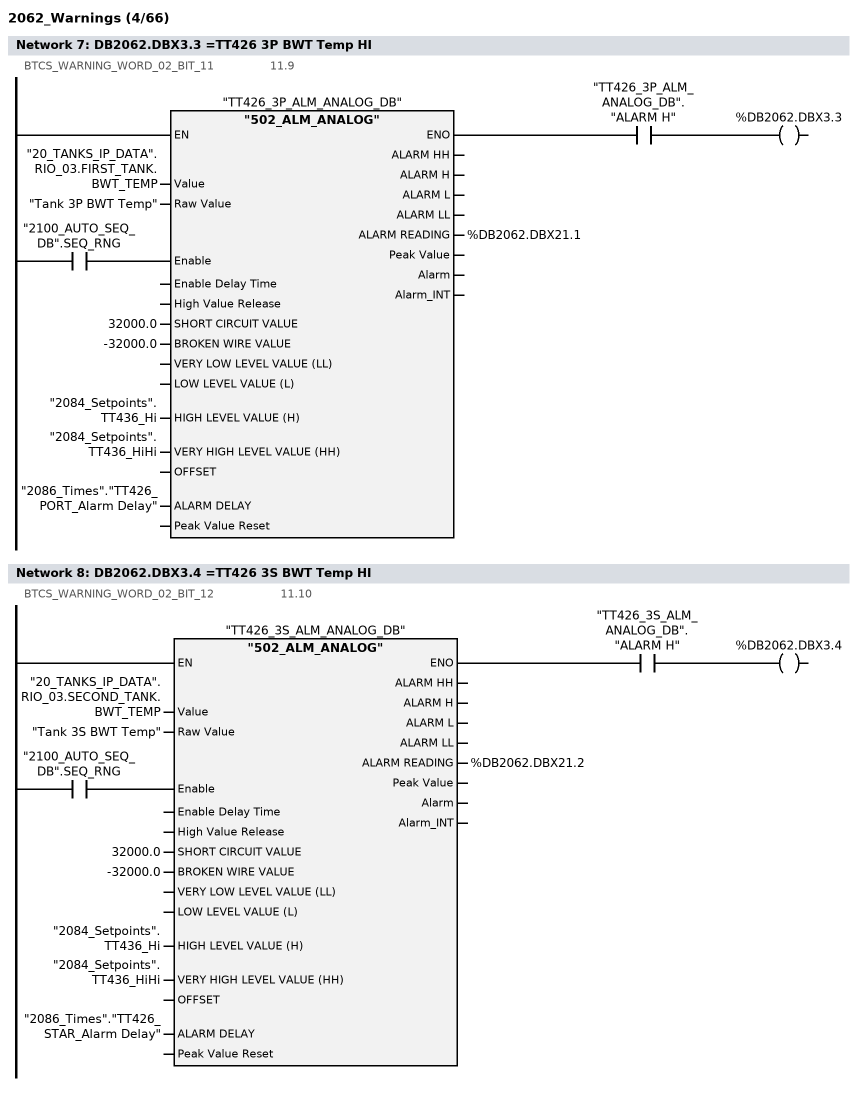
   RUNG wire#powerrail
      "TT426_3P_ALM_ANALOG_DB"(Enable := wire#w1, Value := "20_TANKS_IP_DATA".RIO_03.FIRST_TANK.BWT_TEMP, "Raw Value" := "Tank 3P BWT Temp", "Enable Delay Time" :=, "High Value Release" :=, "SHORT CIRCUIT VALUE" := 32000.0, "BROKEN WIRE VALUE" := -32000.0, "VERY LOW LEVEL VALUE (LL)" :=, "LOW LEVEL VALUE (L)" :=, "HIGH LEVEL VALUE (H)" := "2084_Setpoints".TT436_Hi, "VERY HIGH LEVEL VALUE (HH)" := "2084_Setpoints".TT436_HiHi, OFFSET :=, "ALARM DELAY" := "2086_Times"."TT426_PORT_Alarm Delay", "Peak Value Reset" :=, "ALARM HH" =>, "ALARM H" =>, "ALARM L" =>, "ALARM LL" =>, "ALARM READING" => %DB2062.DBX21.1, "Peak Value" =>, Alarm =>, Alarm_INT =>)
      Contact( "TT426_3P_ALM_ANALOG_DB"."ALARM H" )
      Coil( %DB2062.DBX3.3 )
   END_RUNG
   RUNG wire#powerrail
      Contact( "2100_AUTO_SEQ_DB".SEQ_RNG )
   END_RUNG wire#w1
   // the same network as SCL:
   "TT426_3P_ALM_ANALOG_DB"(Value := "20_TANKS_IP_DATA".RIO_03.FIRST_TANK.BWT_TEMP,   // "502_ALM_ANALOG"
                           "Raw Value" := "Tank 3P BWT Temp",
                           Enable := "2100_AUTO_SEQ_DB".SEQ_RNG,
                           "SHORT CIRCUIT VALUE" := 32000.0,
                           "BROKEN WIRE VALUE" := -32000.0,
                           "HIGH LEVEL VALUE (H)" := "2084_Setpoints".TT436_Hi,
                           "VERY HIGH LEVEL VALUE (HH)" := "2084_Setpoints".TT436_HiHi,
                           "ALARM DELAY" := "2086_Times"."TT426_PORT_Alarm Delay",
                           "ALARM READING" => %DB2062.DBX21.1,
                           ENO => #_w1);
   %DB2062.DBX3.3 := #_w1 AND "TT426_3P_ALM_ANALOG_DB"."ALARM H";
END_REGION

REGION Network 8: DB2062.DBX3.4 =TT426 3S BWT Temp HI
   // BTCS_WARNING_WORD_02_BIT_12                   11.10
   RUNG wire#powerrail
      "TT426_3S_ALM_ANALOG_DB"(Enable := wire#w1, Value := "20_TANKS_IP_DATA".RIO_03.SECOND_TANK.BWT_TEMP, "Raw Value" := "Tank 3S BWT Temp", "Enable Delay Time" :=, "High Value Release" :=, "SHORT CIRCUIT VALUE" := 32000.0, "BROKEN WIRE VALUE" := -32000.0, "VERY LOW LEVEL VALUE (LL)" :=, "LOW LEVEL VALUE (L)" :=, "HIGH LEVEL VALUE (H)" := "2084_Setpoints".TT436_Hi, "VERY HIGH LEVEL VALUE (HH)" := "2084_Setpoints".TT436_HiHi, OFFSET :=, "ALARM DELAY" := "2086_Times"."TT426_STAR_Alarm Delay", "Peak Value Reset" :=, "ALARM HH" =>, "ALARM H" =>, "ALARM L" =>, "ALARM LL" =>, "ALARM READING" => %DB2062.DBX21.2, "Peak Value" =>, Alarm =>, Alarm_INT =>)
      Contact( "TT426_3S_ALM_ANALOG_DB"."ALARM H" )
      Coil( %DB2062.DBX3.4 )
   END_RUNG
   RUNG wire#powerrail
      Contact( "2100_AUTO_SEQ_DB".SEQ_RNG )
   END_RUNG wire#w1
   // the same network as SCL:
   "TT426_3S_ALM_ANALOG_DB"(Value := "20_TANKS_IP_DATA".RIO_03.SECOND_TANK.BWT_TEMP,   // "502_ALM_ANALOG"
                           "Raw Value" := "Tank 3S BWT Temp",
                           Enable := "2100_AUTO_SEQ_DB".SEQ_RNG,
                           "SHORT CIRCUIT VALUE" := 32000.0,
                           "BROKEN WIRE VALUE" := -32000.0,
                           "HIGH LEVEL VALUE (H)" := "2084_Setpoints".TT436_Hi,
                           "VERY HIGH LEVEL VALUE (HH)" := "2084_Setpoints".TT436_HiHi,
                           "ALARM DELAY" := "2086_Times"."TT426_STAR_Alarm Delay",
                           "ALARM READING" => %DB2062.DBX21.2,
                           ENO => #_w1);
   %DB2062.DBX3.4 := #_w1 AND "TT426_3S_ALM_ANALOG_DB"."ALARM H";
END_REGION

REGION Network 9: DB2062.DBX3.5 =TT426 4P BWT Temp HI
   // BTCS_WARNING_WORD_02_BIT_13                     11.11
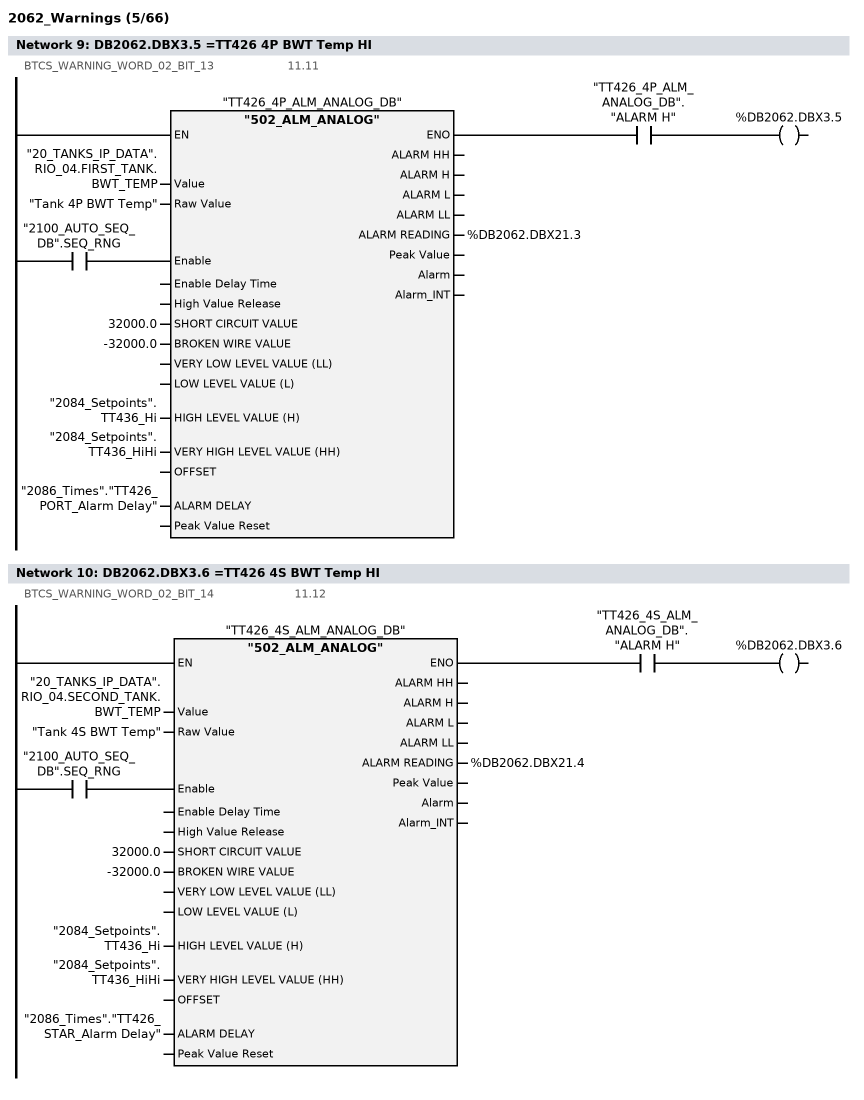
   RUNG wire#powerrail
      "TT426_4P_ALM_ANALOG_DB"(Enable := wire#w1, Value := "20_TANKS_IP_DATA".RIO_04.FIRST_TANK.BWT_TEMP, "Raw Value" := "Tank 4P BWT Temp", "Enable Delay Time" :=, "High Value Release" :=, "SHORT CIRCUIT VALUE" := 32000.0, "BROKEN WIRE VALUE" := -32000.0, "VERY LOW LEVEL VALUE (LL)" :=, "LOW LEVEL VALUE (L)" :=, "HIGH LEVEL VALUE (H)" := "2084_Setpoints".TT436_Hi, "VERY HIGH LEVEL VALUE (HH)" := "2084_Setpoints".TT436_HiHi, OFFSET :=, "ALARM DELAY" := "2086_Times"."TT426_PORT_Alarm Delay", "Peak Value Reset" :=, "ALARM HH" =>, "ALARM H" =>, "ALARM L" =>, "ALARM LL" =>, "ALARM READING" => %DB2062.DBX21.3, "Peak Value" =>, Alarm =>, Alarm_INT =>)
      Contact( "TT426_4P_ALM_ANALOG_DB"."ALARM H" )
      Coil( %DB2062.DBX3.5 )
   END_RUNG
   RUNG wire#powerrail
      Contact( "2100_AUTO_SEQ_DB".SEQ_RNG )
   END_RUNG wire#w1
   // the same network as SCL:
   "TT426_4P_ALM_ANALOG_DB"(Value := "20_TANKS_IP_DATA".RIO_04.FIRST_TANK.BWT_TEMP,   // "502_ALM_ANALOG"
                           "Raw Value" := "Tank 4P BWT Temp",
                           Enable := "2100_AUTO_SEQ_DB".SEQ_RNG,
                           "SHORT CIRCUIT VALUE" := 32000.0,
                           "BROKEN WIRE VALUE" := -32000.0,
                           "HIGH LEVEL VALUE (H)" := "2084_Setpoints".TT436_Hi,
                           "VERY HIGH LEVEL VALUE (HH)" := "2084_Setpoints".TT436_HiHi,
                           "ALARM DELAY" := "2086_Times"."TT426_PORT_Alarm Delay",
                           "ALARM READING" => %DB2062.DBX21.3,
                           ENO => #_w1);
   %DB2062.DBX3.5 := #_w1 AND "TT426_4P_ALM_ANALOG_DB"."ALARM H";
END_REGION

REGION Network 10: DB2062.DBX3.6 =TT426 4S BWT Temp HI
   // BTCS_WARNING_WORD_02_BIT_14                       11.12
   RUNG wire#powerrail
      "TT426_4S_ALM_ANALOG_DB"(Enable := wire#w1, Value := "20_TANKS_IP_DATA".RIO_04.SECOND_TANK.BWT_TEMP, "Raw Value" := "Tank 4S BWT Temp", "Enable Delay Time" :=, "High Value Release" :=, "SHORT CIRCUIT VALUE" := 32000.0, "BROKEN WIRE VALUE" := -32000.0, "VERY LOW LEVEL VALUE (LL)" :=, "LOW LEVEL VALUE (L)" :=, "HIGH LEVEL VALUE (H)" := "2084_Setpoints".TT436_Hi, "VERY HIGH LEVEL VALUE (HH)" := "2084_Setpoints".TT436_HiHi, OFFSET :=, "ALARM DELAY" := "2086_Times"."TT426_STAR_Alarm Delay", "Peak Value Reset" :=, "ALARM HH" =>, "ALARM H" =>, "ALARM L" =>, "ALARM LL" =>, "ALARM READING" => %DB2062.DBX21.4, "Peak Value" =>, Alarm =>, Alarm_INT =>)
      Contact( "TT426_4S_ALM_ANALOG_DB"."ALARM H" )
      Coil( %DB2062.DBX3.6 )
   END_RUNG
   RUNG wire#powerrail
      Contact( "2100_AUTO_SEQ_DB".SEQ_RNG )
   END_RUNG wire#w1
   // the same network as SCL:
   "TT426_4S_ALM_ANALOG_DB"(Value := "20_TANKS_IP_DATA".RIO_04.SECOND_TANK.BWT_TEMP,   // "502_ALM_ANALOG"
                           "Raw Value" := "Tank 4S BWT Temp",
                           Enable := "2100_AUTO_SEQ_DB".SEQ_RNG,
                           "SHORT CIRCUIT VALUE" := 32000.0,
                           "BROKEN WIRE VALUE" := -32000.0,
                           "HIGH LEVEL VALUE (H)" := "2084_Setpoints".TT436_Hi,
                           "VERY HIGH LEVEL VALUE (HH)" := "2084_Setpoints".TT436_HiHi,
                           "ALARM DELAY" := "2086_Times"."TT426_STAR_Alarm Delay",
                           "ALARM READING" => %DB2062.DBX21.4,
                           ENO => #_w1);
   %DB2062.DBX3.6 := #_w1 AND "TT426_4S_ALM_ANALOG_DB"."ALARM H";
END_REGION

REGION Network 11: DB2062.DBX3.7 =TT426 5P BWT Temp HI
   // BTCS_WARNING_WORD_02_BIT_15                        11.13
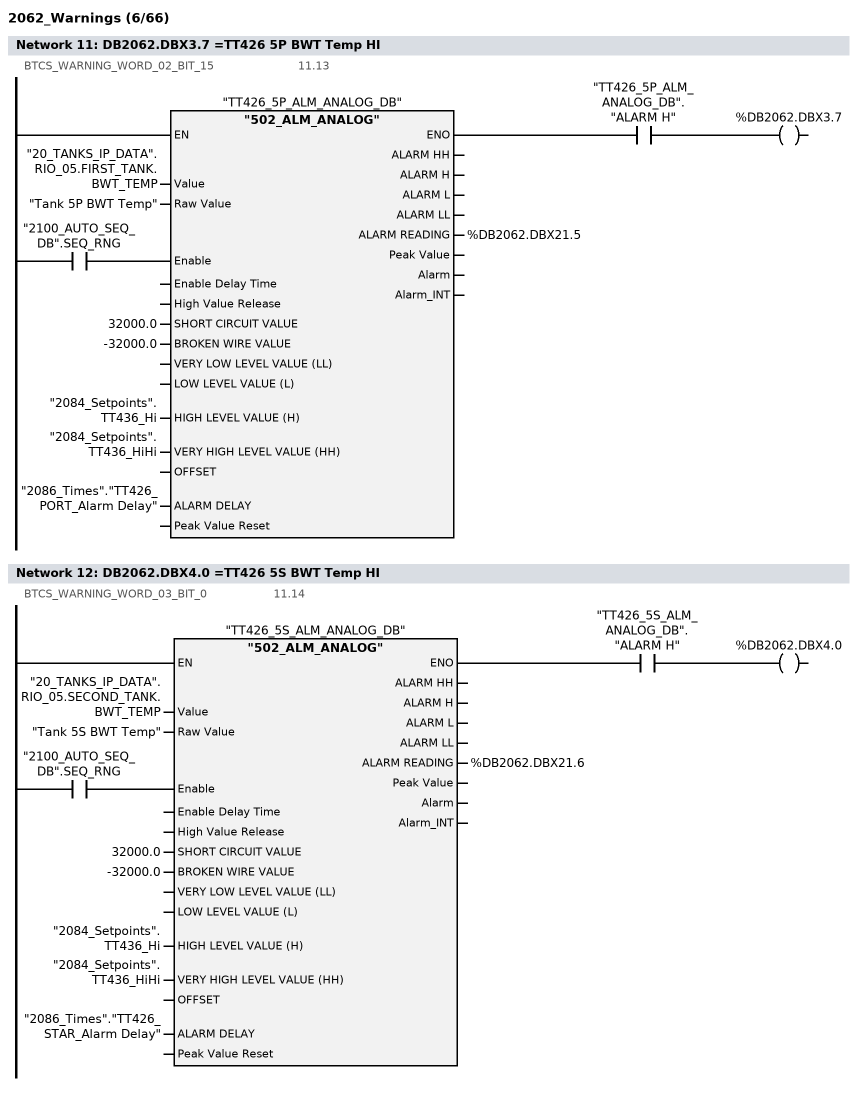
   RUNG wire#powerrail
      "TT426_5P_ALM_ANALOG_DB"(Enable := wire#w1, Value := "20_TANKS_IP_DATA".RIO_05.FIRST_TANK.BWT_TEMP, "Raw Value" := "Tank 5P BWT Temp", "Enable Delay Time" :=, "High Value Release" :=, "SHORT CIRCUIT VALUE" := 32000.0, "BROKEN WIRE VALUE" := -32000.0, "VERY LOW LEVEL VALUE (LL)" :=, "LOW LEVEL VALUE (L)" :=, "HIGH LEVEL VALUE (H)" := "2084_Setpoints".TT436_Hi, "VERY HIGH LEVEL VALUE (HH)" := "2084_Setpoints".TT436_HiHi, OFFSET :=, "ALARM DELAY" := "2086_Times"."TT426_PORT_Alarm Delay", "Peak Value Reset" :=, "ALARM HH" =>, "ALARM H" =>, "ALARM L" =>, "ALARM LL" =>, "ALARM READING" => %DB2062.DBX21.5, "Peak Value" =>, Alarm =>, Alarm_INT =>)
      Contact( "TT426_5P_ALM_ANALOG_DB"."ALARM H" )
      Coil( %DB2062.DBX3.7 )
   END_RUNG
   RUNG wire#powerrail
      Contact( "2100_AUTO_SEQ_DB".SEQ_RNG )
   END_RUNG wire#w1
   // the same network as SCL:
   "TT426_5P_ALM_ANALOG_DB"(Value := "20_TANKS_IP_DATA".RIO_05.FIRST_TANK.BWT_TEMP,   // "502_ALM_ANALOG"
                           "Raw Value" := "Tank 5P BWT Temp",
                           Enable := "2100_AUTO_SEQ_DB".SEQ_RNG,
                           "SHORT CIRCUIT VALUE" := 32000.0,
                           "BROKEN WIRE VALUE" := -32000.0,
                           "HIGH LEVEL VALUE (H)" := "2084_Setpoints".TT436_Hi,
                           "VERY HIGH LEVEL VALUE (HH)" := "2084_Setpoints".TT436_HiHi,
                           "ALARM DELAY" := "2086_Times"."TT426_PORT_Alarm Delay",
                           "ALARM READING" => %DB2062.DBX21.5,
                           ENO => #_w1);
   %DB2062.DBX3.7 := #_w1 AND "TT426_5P_ALM_ANALOG_DB"."ALARM H";
END_REGION

REGION Network 12: DB2062.DBX4.0 =TT426 5S BWT Temp HI
   // BTCS_WARNING_WORD_03_BIT_0                   11.14
   RUNG wire#powerrail
      "TT426_5S_ALM_ANALOG_DB"(Enable := wire#w1, Value := "20_TANKS_IP_DATA".RIO_05.SECOND_TANK.BWT_TEMP, "Raw Value" := "Tank 5S BWT Temp", "Enable Delay Time" :=, "High Value Release" :=, "SHORT CIRCUIT VALUE" := 32000.0, "BROKEN WIRE VALUE" := -32000.0, "VERY LOW LEVEL VALUE (LL)" :=, "LOW LEVEL VALUE (L)" :=, "HIGH LEVEL VALUE (H)" := "2084_Setpoints".TT436_Hi, "VERY HIGH LEVEL VALUE (HH)" := "2084_Setpoints".TT436_HiHi, OFFSET :=, "ALARM DELAY" := "2086_Times"."TT426_STAR_Alarm Delay", "Peak Value Reset" :=, "ALARM HH" =>, "ALARM H" =>, "ALARM L" =>, "ALARM LL" =>, "ALARM READING" => %DB2062.DBX21.6, "Peak Value" =>, Alarm =>, Alarm_INT =>)
      Contact( "TT426_5S_ALM_ANALOG_DB"."ALARM H" )
      Coil( %DB2062.DBX4.0 )
   END_RUNG
   RUNG wire#powerrail
      Contact( "2100_AUTO_SEQ_DB".SEQ_RNG )
   END_RUNG wire#w1
   // the same network as SCL:
   "TT426_5S_ALM_ANALOG_DB"(Value := "20_TANKS_IP_DATA".RIO_05.SECOND_TANK.BWT_TEMP,   // "502_ALM_ANALOG"
                           "Raw Value" := "Tank 5S BWT Temp",
                           Enable := "2100_AUTO_SEQ_DB".SEQ_RNG,
                           "SHORT CIRCUIT VALUE" := 32000.0,
                           "BROKEN WIRE VALUE" := -32000.0,
                           "HIGH LEVEL VALUE (H)" := "2084_Setpoints".TT436_Hi,
                           "VERY HIGH LEVEL VALUE (HH)" := "2084_Setpoints".TT436_HiHi,
                           "ALARM DELAY" := "2086_Times"."TT426_STAR_Alarm Delay",
                           "ALARM READING" => %DB2062.DBX21.6,
                           ENO => #_w1);
   %DB2062.DBX4.0 := #_w1 AND "TT426_5S_ALM_ANALOG_DB"."ALARM H";
END_REGION

REGION Network 13: DB2062.DBX4.1 =TT426 6P BWT Temp HI
   // BTCS_WARNING_WORD_03_BIT_1                           11.15
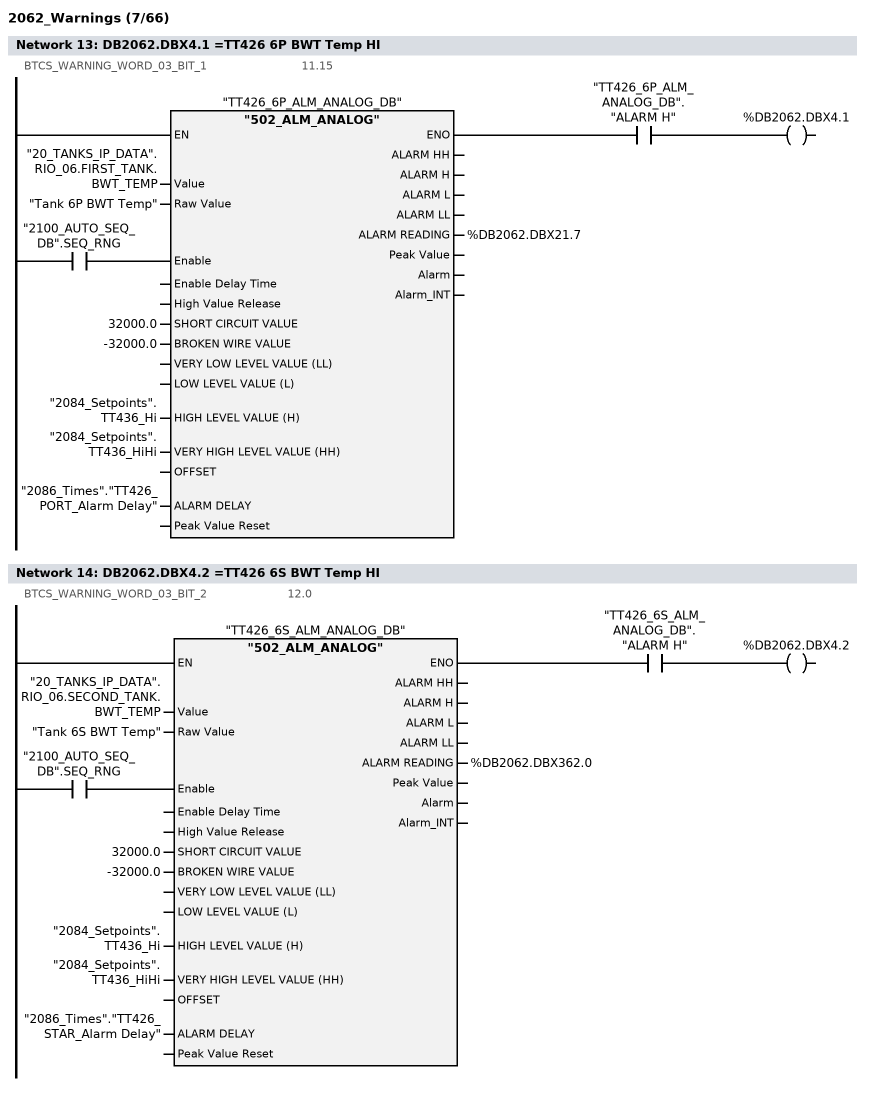
   RUNG wire#powerrail
      "TT426_6P_ALM_ANALOG_DB"(Enable := wire#w1, Value := "20_TANKS_IP_DATA".RIO_06.FIRST_TANK.BWT_TEMP, "Raw Value" := "Tank 6P BWT Temp", "Enable Delay Time" :=, "High Value Release" :=, "SHORT CIRCUIT VALUE" := 32000.0, "BROKEN WIRE VALUE" := -32000.0, "VERY LOW LEVEL VALUE (LL)" :=, "LOW LEVEL VALUE (L)" :=, "HIGH LEVEL VALUE (H)" := "2084_Setpoints".TT436_Hi, "VERY HIGH LEVEL VALUE (HH)" := "2084_Setpoints".TT436_HiHi, OFFSET :=, "ALARM DELAY" := "2086_Times"."TT426_PORT_Alarm Delay", "Peak Value Reset" :=, "ALARM HH" =>, "ALARM H" =>, "ALARM L" =>, "ALARM LL" =>, "ALARM READING" => %DB2062.DBX21.7, "Peak Value" =>, Alarm =>, Alarm_INT =>)
      Contact( "TT426_6P_ALM_ANALOG_DB"."ALARM H" )
      Coil( %DB2062.DBX4.1 )
   END_RUNG
   RUNG wire#powerrail
      Contact( "2100_AUTO_SEQ_DB".SEQ_RNG )
   END_RUNG wire#w1
   // the same network as SCL:
   "TT426_6P_ALM_ANALOG_DB"(Value := "20_TANKS_IP_DATA".RIO_06.FIRST_TANK.BWT_TEMP,   // "502_ALM_ANALOG"
                           "Raw Value" := "Tank 6P BWT Temp",
                           Enable := "2100_AUTO_SEQ_DB".SEQ_RNG,
                           "SHORT CIRCUIT VALUE" := 32000.0,
                           "BROKEN WIRE VALUE" := -32000.0,
                           "HIGH LEVEL VALUE (H)" := "2084_Setpoints".TT436_Hi,
                           "VERY HIGH LEVEL VALUE (HH)" := "2084_Setpoints".TT436_HiHi,
                           "ALARM DELAY" := "2086_Times"."TT426_PORT_Alarm Delay",
                           "ALARM READING" => %DB2062.DBX21.7,
                           ENO => #_w1);
   %DB2062.DBX4.1 := #_w1 AND "TT426_6P_ALM_ANALOG_DB"."ALARM H";
END_REGION

REGION Network 14: DB2062.DBX4.2 =TT426 6S BWT Temp HI
   // BTCS_WARNING_WORD_03_BIT_2                       12.0
   RUNG wire#powerrail
      "TT426_6S_ALM_ANALOG_DB"(Enable := wire#w1, Value := "20_TANKS_IP_DATA".RIO_06.SECOND_TANK.BWT_TEMP, "Raw Value" := "Tank 6S BWT Temp", "Enable Delay Time" :=, "High Value Release" :=, "SHORT CIRCUIT VALUE" := 32000.0, "BROKEN WIRE VALUE" := -32000.0, "VERY LOW LEVEL VALUE (LL)" :=, "LOW LEVEL VALUE (L)" :=, "HIGH LEVEL VALUE (H)" := "2084_Setpoints".TT436_Hi, "VERY HIGH LEVEL VALUE (HH)" := "2084_Setpoints".TT436_HiHi, OFFSET :=, "ALARM DELAY" := "2086_Times"."TT426_STAR_Alarm Delay", "Peak Value Reset" :=, "ALARM HH" =>, "ALARM H" =>, "ALARM L" =>, "ALARM LL" =>, "ALARM READING" => %DB2062.DBX362.0, "Peak Value" =>, Alarm =>, Alarm_INT =>)
      Contact( "TT426_6S_ALM_ANALOG_DB"."ALARM H" )
      Coil( %DB2062.DBX4.2 )
   END_RUNG
   RUNG wire#powerrail
      Contact( "2100_AUTO_SEQ_DB".SEQ_RNG )
   END_RUNG wire#w1
   // the same network as SCL:
   "TT426_6S_ALM_ANALOG_DB"(Value := "20_TANKS_IP_DATA".RIO_06.SECOND_TANK.BWT_TEMP,   // "502_ALM_ANALOG"
                           "Raw Value" := "Tank 6S BWT Temp",
                           Enable := "2100_AUTO_SEQ_DB".SEQ_RNG,
                           "SHORT CIRCUIT VALUE" := 32000.0,
                           "BROKEN WIRE VALUE" := -32000.0,
                           "HIGH LEVEL VALUE (H)" := "2084_Setpoints".TT436_Hi,
                           "VERY HIGH LEVEL VALUE (HH)" := "2084_Setpoints".TT436_HiHi,
                           "ALARM DELAY" := "2086_Times"."TT426_STAR_Alarm Delay",
                           "ALARM READING" => %DB2062.DBX362.0,
                           ENO => #_w1);
   %DB2062.DBX4.2 := #_w1 AND "TT426_6S_ALM_ANALOG_DB"."ALARM H";
END_REGION

REGION Network 15: DB2062.DBX4.3 =TT426 APT BWT Temp HI
   // BTCS_WARNING_WORD_03_BIT_3                                 12.1
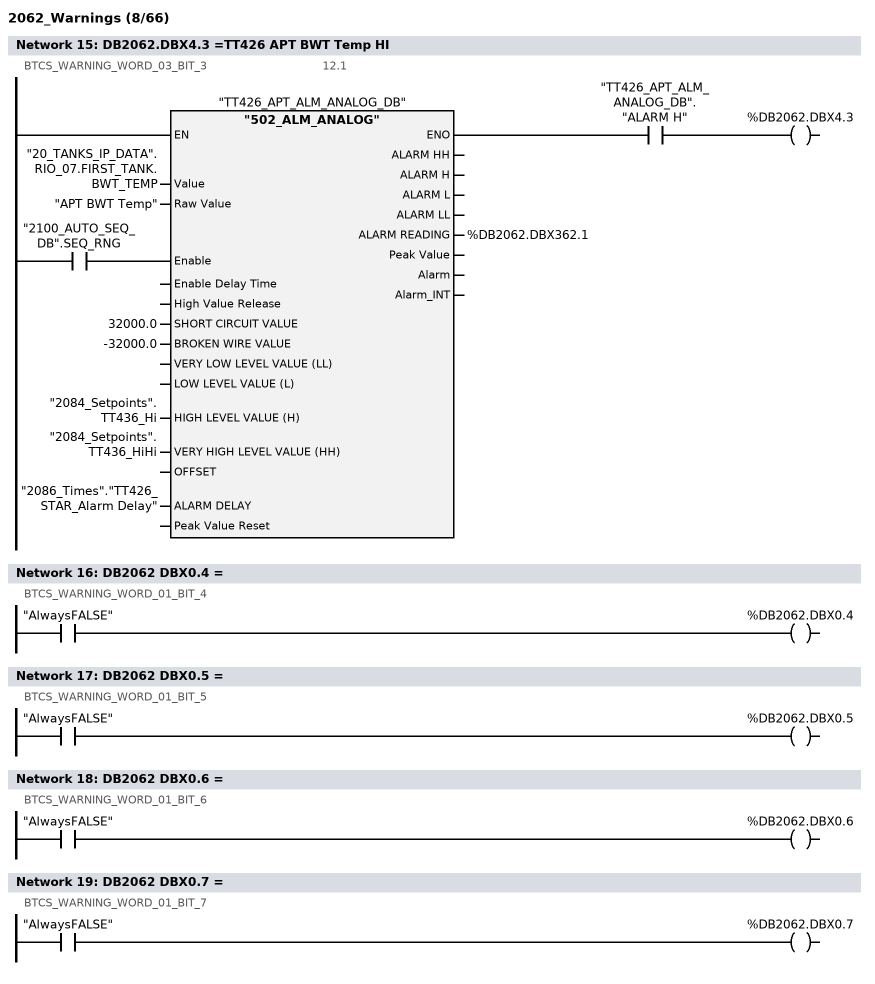
   RUNG wire#powerrail
      "TT426_APT_ALM_ANALOG_DB"(Enable := wire#w1, Value := "20_TANKS_IP_DATA".RIO_07.FIRST_TANK.BWT_TEMP, "Raw Value" := "APT BWT Temp", "Enable Delay Time" :=, "High Value Release" :=, "SHORT CIRCUIT VALUE" := 32000.0, "BROKEN WIRE VALUE" := -32000.0, "VERY LOW LEVEL VALUE (LL)" :=, "LOW LEVEL VALUE (L)" :=, "HIGH LEVEL VALUE (H)" := "2084_Setpoints".TT436_Hi, "VERY HIGH LEVEL VALUE (HH)" := "2084_Setpoints".TT436_HiHi, OFFSET :=, "ALARM DELAY" := "2086_Times"."TT426_STAR_Alarm Delay", "Peak Value Reset" :=, "ALARM HH" =>, "ALARM H" =>, "ALARM L" =>, "ALARM LL" =>, "ALARM READING" => %DB2062.DBX362.1, "Peak Value" =>, Alarm =>, Alarm_INT =>)
      Contact( "TT426_APT_ALM_ANALOG_DB"."ALARM H" )
      Coil( %DB2062.DBX4.3 )
   END_RUNG
   RUNG wire#powerrail
      Contact( "2100_AUTO_SEQ_DB".SEQ_RNG )
   END_RUNG wire#w1
   // the same network as SCL:
   "TT426_APT_ALM_ANALOG_DB"(Value := "20_TANKS_IP_DATA".RIO_07.FIRST_TANK.BWT_TEMP,   // "502_ALM_ANALOG"
                           "Raw Value" := "APT BWT Temp",
                           Enable := "2100_AUTO_SEQ_DB".SEQ_RNG,
                           "SHORT CIRCUIT VALUE" := 32000.0,
                           "BROKEN WIRE VALUE" := -32000.0,
                           "HIGH LEVEL VALUE (H)" := "2084_Setpoints".TT436_Hi,
                           "VERY HIGH LEVEL VALUE (HH)" := "2084_Setpoints".TT436_HiHi,
                           "ALARM DELAY" := "2086_Times"."TT426_STAR_Alarm Delay",
                           "ALARM READING" => %DB2062.DBX362.1,
                           ENO => #_w1);
   %DB2062.DBX4.3 := #_w1 AND "TT426_APT_ALM_ANALOG_DB"."ALARM H";
END_REGION

REGION Network 16: DB2062 DBX0.4 =
   // BTCS_WARNING_WORD_01_BIT_4
   RUNG wire#powerrail
      Contact( "AlwaysFALSE" )
      Coil( %DB2062.DBX0.4 )
   END_RUNG
   // the same network as SCL:
   %DB2062.DBX0.4 := "AlwaysFALSE";
END_REGION

REGION Network 17: DB2062 DBX0.5 =
   // BTCS_WARNING_WORD_01_BIT_5
   RUNG wire#powerrail
      Contact( "AlwaysFALSE" )
      Coil( %DB2062.DBX0.5 )
   END_RUNG
   // the same network as SCL:
   %DB2062.DBX0.5 := "AlwaysFALSE";
END_REGION

REGION Network 18: DB2062 DBX0.6 =
   // BTCS_WARNING_WORD_01_BIT_6
   RUNG wire#powerrail
      Contact( "AlwaysFALSE" )
      Coil( %DB2062.DBX0.6 )
   END_RUNG
   // the same network as SCL:
   %DB2062.DBX0.6 := "AlwaysFALSE";
END_REGION

REGION Network 19: DB2062 DBX0.7 =
   // BTCS_WARNING_WORD_01_BIT_7
   RUNG wire#powerrail
      Contact( "AlwaysFALSE" )
      Coil( %DB2062.DBX0.7 )
   END_RUNG
   // the same network as SCL:
   %DB2062.DBX0.7 := "AlwaysFALSE";
END_REGION

REGION Network 20: DB2062.DBX5.0 = FIT418 FPT USD Flow LO / DB2062.DBX5.1 = FIT418 FPT USD Flow HI
   // BTCS_WARNING_WORD_03_BIT_8/9                    12.2
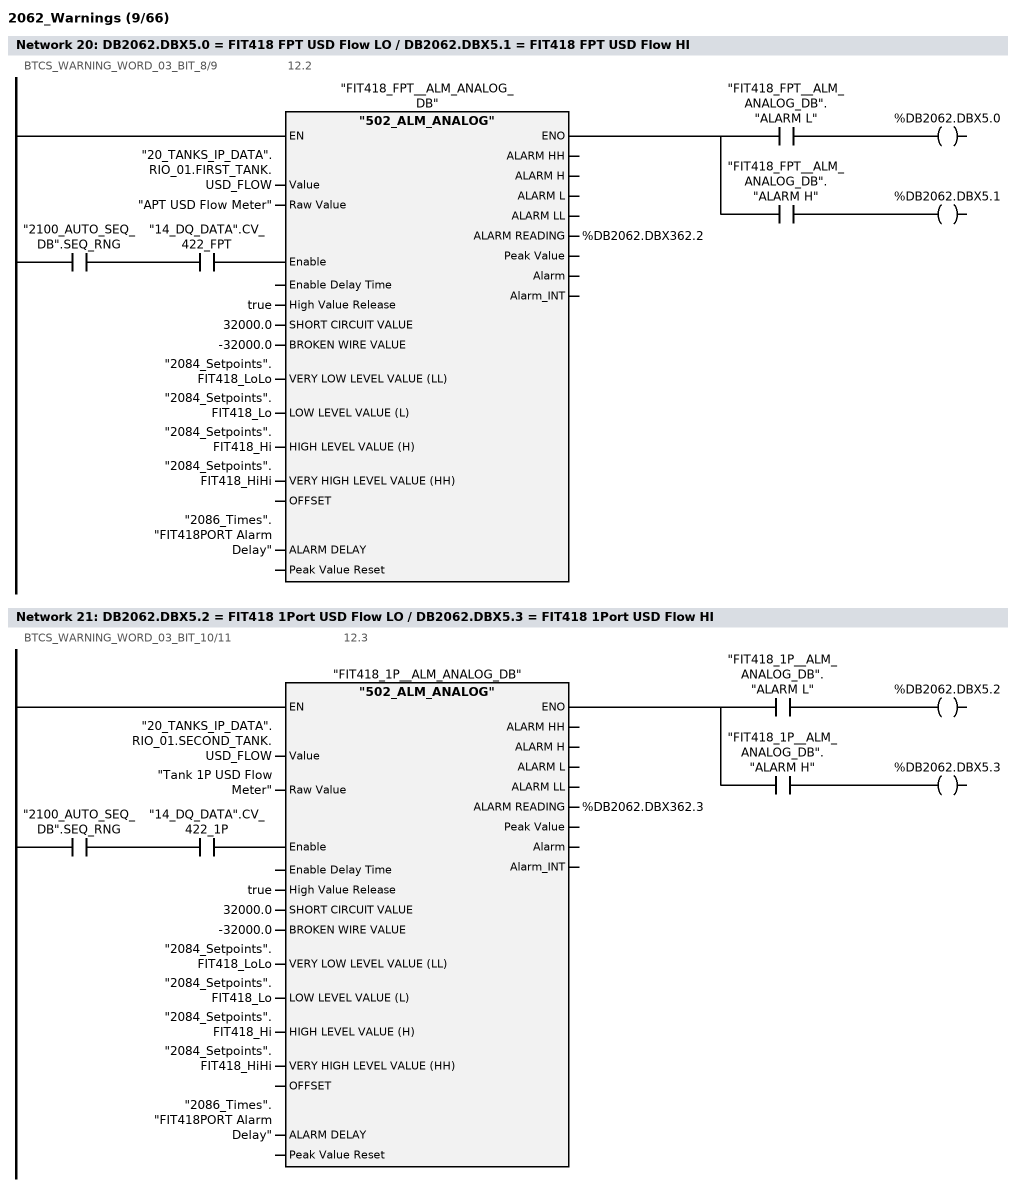
   RUNG wire#powerrail
      "FIT418_FPT__ALM_ANALOG_DB"(Enable := wire#w1, Value := "20_TANKS_IP_DATA".RIO_01.FIRST_TANK.USD_FLOW, "Raw Value" := "APT USD Flow Meter", "Enable Delay Time" :=, "High Value Release" := true, "SHORT CIRCUIT VALUE" := 32000.0, "BROKEN WIRE VALUE" := -32000.0, "VERY LOW LEVEL VALUE (LL)" := "2084_Setpoints".FIT418_LoLo, "LOW LEVEL VALUE (L)" := "2084_Setpoints".FIT418_Lo, "HIGH LEVEL VALUE (H)" := "2084_Setpoints".FIT418_Hi, "VERY HIGH LEVEL VALUE (HH)" := "2084_Setpoints".FIT418_HiHi, OFFSET :=, "ALARM DELAY" := "2086_Times"."FIT418PORT Alarm Delay", "Peak Value Reset" :=, "ALARM HH" =>, "ALARM H" =>, "ALARM L" =>, "ALARM LL" =>, "ALARM READING" => %DB2062.DBX362.2, "Peak Value" =>, Alarm =>, Alarm_INT =>)
      wire#w2
      Contact( "FIT418_FPT__ALM_ANALOG_DB"."ALARM L" )
      Coil( %DB2062.DBX5.0 )
   END_RUNG
   RUNG wire#powerrail
      Contact( "2100_AUTO_SEQ_DB".SEQ_RNG )
      Contact( "14_DQ_DATA".CV_422_FPT )
   END_RUNG wire#w1
   RUNG wire#w2
      Contact( "FIT418_FPT__ALM_ANALOG_DB"."ALARM H" )
      Coil( %DB2062.DBX5.1 )
   END_RUNG
   // the same network as SCL:
   "FIT418_FPT__ALM_ANALOG_DB"(Value := "20_TANKS_IP_DATA".RIO_01.FIRST_TANK.USD_FLOW,   // "502_ALM_ANALOG"
                           "Raw Value" := "APT USD Flow Meter",
                           Enable := "2100_AUTO_SEQ_DB".SEQ_RNG AND "14_DQ_DATA".CV_422_FPT,
                           "High Value Release" := true,
                           "SHORT CIRCUIT VALUE" := 32000.0,
                           "BROKEN WIRE VALUE" := -32000.0,
                           "VERY LOW LEVEL VALUE (LL)" := "2084_Setpoints".FIT418_LoLo,
                           "LOW LEVEL VALUE (L)" := "2084_Setpoints".FIT418_Lo,
                           "HIGH LEVEL VALUE (H)" := "2084_Setpoints".FIT418_Hi,
                           "VERY HIGH LEVEL VALUE (HH)" := "2084_Setpoints".FIT418_HiHi,
                           "ALARM DELAY" := "2086_Times"."FIT418PORT Alarm Delay",
                           "ALARM READING" => %DB2062.DBX362.2,
                           ENO => #_w1);
   %DB2062.DBX5.0 := #_w1 AND "FIT418_FPT__ALM_ANALOG_DB"."ALARM L";
   %DB2062.DBX5.1 := #_w1 AND "FIT418_FPT__ALM_ANALOG_DB"."ALARM H";
END_REGION

REGION Network 21: DB2062.DBX5.2 = FIT418 1Port USD Flow LO / DB2062.DBX5.3 = FIT418 1Port USD Flow HI
   // BTCS_WARNING_WORD_03_BIT_10/11                                12.3
   RUNG wire#powerrail
      "FIT418_1P__ALM_ANALOG_DB"(Enable := wire#w1, Value := "20_TANKS_IP_DATA".RIO_01.SECOND_TANK.USD_FLOW, "Raw Value" := "Tank 1P USD Flow Meter", "Enable Delay Time" :=, "High Value Release" := true, "SHORT CIRCUIT VALUE" := 32000.0, "BROKEN WIRE VALUE" := -32000.0, "VERY LOW LEVEL VALUE (LL)" := "2084_Setpoints".FIT418_LoLo, "LOW LEVEL VALUE (L)" := "2084_Setpoints".FIT418_Lo, "HIGH LEVEL VALUE (H)" := "2084_Setpoints".FIT418_Hi, "VERY HIGH LEVEL VALUE (HH)" := "2084_Setpoints".FIT418_HiHi, OFFSET :=, "ALARM DELAY" := "2086_Times"."FIT418PORT Alarm Delay", "Peak Value Reset" :=, "ALARM HH" =>, "ALARM H" =>, "ALARM L" =>, "ALARM LL" =>, "ALARM READING" => %DB2062.DBX362.3, "Peak Value" =>, Alarm =>, Alarm_INT =>)
      wire#w2
      Contact( "FIT418_1P__ALM_ANALOG_DB"."ALARM L" )
      Coil( %DB2062.DBX5.2 )
   END_RUNG
   RUNG wire#powerrail
      Contact( "2100_AUTO_SEQ_DB".SEQ_RNG )
      Contact( "14_DQ_DATA".CV_422_1P )
   END_RUNG wire#w1
   RUNG wire#w2
      Contact( "FIT418_1P__ALM_ANALOG_DB"."ALARM H" )
      Coil( %DB2062.DBX5.3 )
   END_RUNG
   // the same network as SCL:
   "FIT418_1P__ALM_ANALOG_DB"(Value := "20_TANKS_IP_DATA".RIO_01.SECOND_TANK.USD_FLOW,   // "502_ALM_ANALOG"
                           "Raw Value" := "Tank 1P USD Flow Meter",
                           Enable := "2100_AUTO_SEQ_DB".SEQ_RNG AND "14_DQ_DATA".CV_422_1P,
                           "High Value Release" := true,
                           "SHORT CIRCUIT VALUE" := 32000.0,
                           "BROKEN WIRE VALUE" := -32000.0,
                           "VERY LOW LEVEL VALUE (LL)" := "2084_Setpoints".FIT418_LoLo,
                           "LOW LEVEL VALUE (L)" := "2084_Setpoints".FIT418_Lo,
                           "HIGH LEVEL VALUE (H)" := "2084_Setpoints".FIT418_Hi,
                           "VERY HIGH LEVEL VALUE (HH)" := "2084_Setpoints".FIT418_HiHi,
                           "ALARM DELAY" := "2086_Times"."FIT418PORT Alarm Delay",
                           "ALARM READING" => %DB2062.DBX362.3,
                           ENO => #_w1);
   %DB2062.DBX5.2 := #_w1 AND "FIT418_1P__ALM_ANALOG_DB"."ALARM L";
   %DB2062.DBX5.3 := #_w1 AND "FIT418_1P__ALM_ANALOG_DB"."ALARM H";
END_REGION

REGION Network 22: DB2062.DBX5.4 = FIT417 1Star USD Flow LO / DB2062.DBX5.5 = FIT417 1Star USD Flow HI
   // BTCS_WARNING_WORD_03_BIT_12/13                        12.4
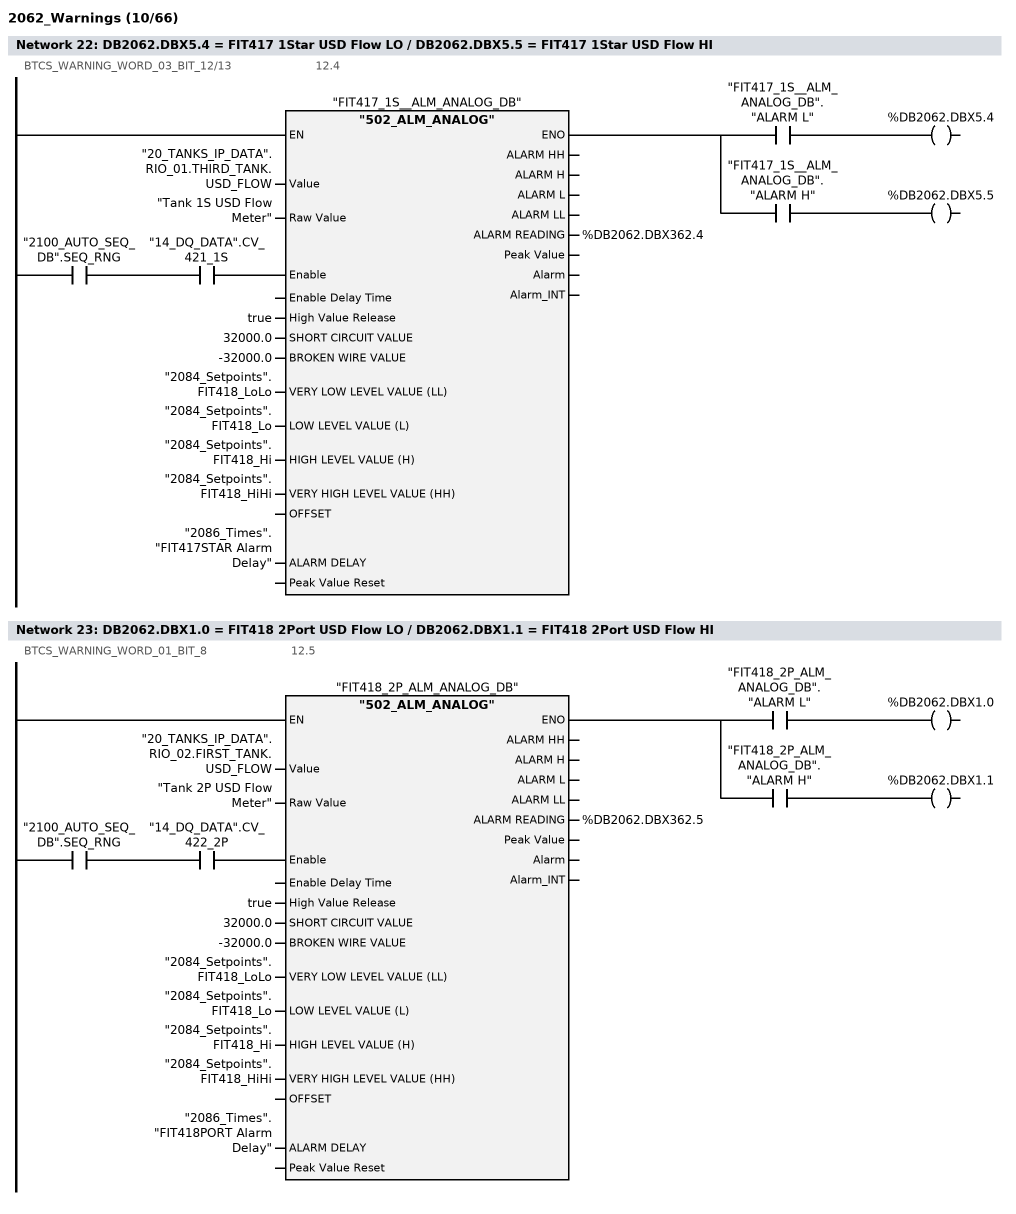
   RUNG wire#powerrail
      "FIT417_1S__ALM_ANALOG_DB"(Enable := wire#w1, Value := "20_TANKS_IP_DATA".RIO_01.THIRD_TANK.USD_FLOW, "Raw Value" := "Tank 1S USD Flow Meter", "Enable Delay Time" :=, "High Value Release" := true, "SHORT CIRCUIT VALUE" := 32000.0, "BROKEN WIRE VALUE" := -32000.0, "VERY LOW LEVEL VALUE (LL)" := "2084_Setpoints".FIT418_LoLo, "LOW LEVEL VALUE (L)" := "2084_Setpoints".FIT418_Lo, "HIGH LEVEL VALUE (H)" := "2084_Setpoints".FIT418_Hi, "VERY HIGH LEVEL VALUE (HH)" := "2084_Setpoints".FIT418_HiHi, OFFSET :=, "ALARM DELAY" := "2086_Times"."FIT417STAR Alarm Delay", "Peak Value Reset" :=, "ALARM HH" =>, "ALARM H" =>, "ALARM L" =>, "ALARM LL" =>, "ALARM READING" => %DB2062.DBX362.4, "Peak Value" =>, Alarm =>, Alarm_INT =>)
      wire#w2
      Contact( "FIT417_1S__ALM_ANALOG_DB"."ALARM L" )
      Coil( %DB2062.DBX5.4 )
   END_RUNG
   RUNG wire#powerrail
      Contact( "2100_AUTO_SEQ_DB".SEQ_RNG )
      Contact( "14_DQ_DATA".CV_421_1S )
   END_RUNG wire#w1
   RUNG wire#w2
      Contact( "FIT417_1S__ALM_ANALOG_DB"."ALARM H" )
      Coil( %DB2062.DBX5.5 )
   END_RUNG
   // the same network as SCL:
   "FIT417_1S__ALM_ANALOG_DB"(Value := "20_TANKS_IP_DATA".RIO_01.THIRD_TANK.USD_FLOW,   // "502_ALM_ANALOG"
                           "Raw Value" := "Tank 1S USD Flow Meter",
                           Enable := "2100_AUTO_SEQ_DB".SEQ_RNG AND "14_DQ_DATA".CV_421_1S,
                           "High Value Release" := true,
                           "SHORT CIRCUIT VALUE" := 32000.0,
                           "BROKEN WIRE VALUE" := -32000.0,
                           "VERY LOW LEVEL VALUE (LL)" := "2084_Setpoints".FIT418_LoLo,
                           "LOW LEVEL VALUE (L)" := "2084_Setpoints".FIT418_Lo,
                           "HIGH LEVEL VALUE (H)" := "2084_Setpoints".FIT418_Hi,
                           "VERY HIGH LEVEL VALUE (HH)" := "2084_Setpoints".FIT418_HiHi,
                           "ALARM DELAY" := "2086_Times"."FIT417STAR Alarm Delay",
                           "ALARM READING" => %DB2062.DBX362.4,
                           ENO => #_w1);
   %DB2062.DBX5.4 := #_w1 AND "FIT417_1S__ALM_ANALOG_DB"."ALARM L";
   %DB2062.DBX5.5 := #_w1 AND "FIT417_1S__ALM_ANALOG_DB"."ALARM H";
END_REGION

REGION Network 23: DB2062.DBX1.0 = FIT418 2Port USD Flow LO / DB2062.DBX1.1 = FIT418 2Port USD Flow HI
   // BTCS_WARNING_WORD_01_BIT_8                        12.5
   RUNG wire#powerrail
      "FIT418_2P_ALM_ANALOG_DB"(Enable := wire#w1, Value := "20_TANKS_IP_DATA".RIO_02.FIRST_TANK.USD_FLOW, "Raw Value" := "Tank 2P USD Flow Meter", "Enable Delay Time" :=, "High Value Release" := true, "SHORT CIRCUIT VALUE" := 32000.0, "BROKEN WIRE VALUE" := -32000.0, "VERY LOW LEVEL VALUE (LL)" := "2084_Setpoints".FIT418_LoLo, "LOW LEVEL VALUE (L)" := "2084_Setpoints".FIT418_Lo, "HIGH LEVEL VALUE (H)" := "2084_Setpoints".FIT418_Hi, "VERY HIGH LEVEL VALUE (HH)" := "2084_Setpoints".FIT418_HiHi, OFFSET :=, "ALARM DELAY" := "2086_Times"."FIT418PORT Alarm Delay", "Peak Value Reset" :=, "ALARM HH" =>, "ALARM H" =>, "ALARM L" =>, "ALARM LL" =>, "ALARM READING" => %DB2062.DBX362.5, "Peak Value" =>, Alarm =>, Alarm_INT =>)
      wire#w2
      Contact( "FIT418_2P_ALM_ANALOG_DB"."ALARM L" )
      Coil( %DB2062.DBX1.0 )
   END_RUNG
   RUNG wire#powerrail
      Contact( "2100_AUTO_SEQ_DB".SEQ_RNG )
      Contact( "14_DQ_DATA".CV_422_2P )
   END_RUNG wire#w1
   RUNG wire#w2
      Contact( "FIT418_2P_ALM_ANALOG_DB"."ALARM H" )
      Coil( %DB2062.DBX1.1 )
   END_RUNG
   // the same network as SCL:
   "FIT418_2P_ALM_ANALOG_DB"(Value := "20_TANKS_IP_DATA".RIO_02.FIRST_TANK.USD_FLOW,   // "502_ALM_ANALOG"
                           "Raw Value" := "Tank 2P USD Flow Meter",
                           Enable := "2100_AUTO_SEQ_DB".SEQ_RNG AND "14_DQ_DATA".CV_422_2P,
                           "High Value Release" := true,
                           "SHORT CIRCUIT VALUE" := 32000.0,
                           "BROKEN WIRE VALUE" := -32000.0,
                           "VERY LOW LEVEL VALUE (LL)" := "2084_Setpoints".FIT418_LoLo,
                           "LOW LEVEL VALUE (L)" := "2084_Setpoints".FIT418_Lo,
                           "HIGH LEVEL VALUE (H)" := "2084_Setpoints".FIT418_Hi,
                           "VERY HIGH LEVEL VALUE (HH)" := "2084_Setpoints".FIT418_HiHi,
                           "ALARM DELAY" := "2086_Times"."FIT418PORT Alarm Delay",
                           "ALARM READING" => %DB2062.DBX362.5,
                           ENO => #_w1);
   %DB2062.DBX1.0 := #_w1 AND "FIT418_2P_ALM_ANALOG_DB"."ALARM L";
   %DB2062.DBX1.1 := #_w1 AND "FIT418_2P_ALM_ANALOG_DB"."ALARM H";
END_REGION

REGION Network 24: DB2062.DBX1.4 = FIT417 2Starboard USD Flow LO / DB2062.DBX1.5 = FIT417 2Starboard USD Flow HI
   // BTCS_WARNING_WORD_01_BIT_12                          12.6